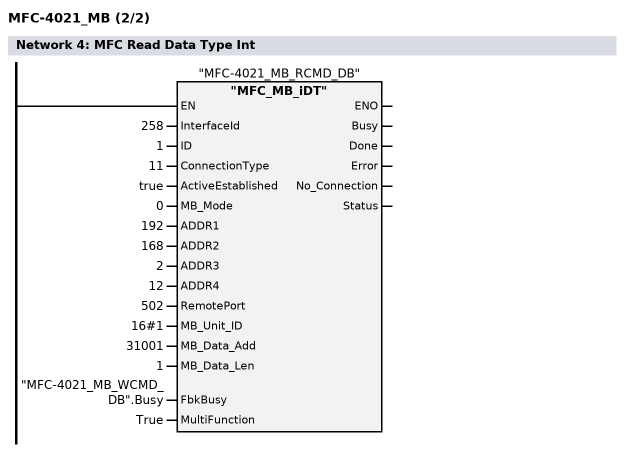
   RUNG wire#powerrail
      "MFC-4021_MB_RCMD_DB"(InterfaceId := 258, ID := 1, ConnectionType := 11, ActiveEstablished := true, MB_Mode := 0, ADDR1 := 192, ADDR2 := 168, ADDR3 := 2, ADDR4 := 12, RemotePort := 502, MB_Unit_ID := 16#1, MB_Data_Add := 31001, MB_Data_Len := 1, FbkBusy := "MFC-4021_MB_WCMD_DB".Busy, MultiFunction := True, Busy =>, Done =>, Error =>, No_Connection =>, Status =>)
   END_RUNG
   // the same network as SCL:
   "MFC-4021_MB_RCMD_DB"(InterfaceId := 258,   // "MFC_MB_iDT"
                         ID := 1,
                         ConnectionType := 11,
                         ActiveEstablished := true,
                         MB_Mode := 0,
                         ADDR1 := 192,
                         ADDR2 := 168,
                         ADDR3 := 2,
                         ADDR4 := 12,
                         RemotePort := 502,
                         MB_Unit_ID := 16#1,
                         MB_Data_Add := 31001,
                         MB_Data_Len := 1,
                         FbkBusy := "MFC-4021_MB_WCMD_DB".Busy,
                         MultiFunction := True);
END_REGION
END_FUNCTION

// folder: Outside Comms/ModBus Comms/MFCs/MFC-4024

FUNCTION "MFC-4024_MB" : Void   // FC78, LAD
{ S7_Optimized_Access := 'TRUE' }
VERSION : 0.1
BEGIN

REGION Network 1: MFC Read Data Type Real
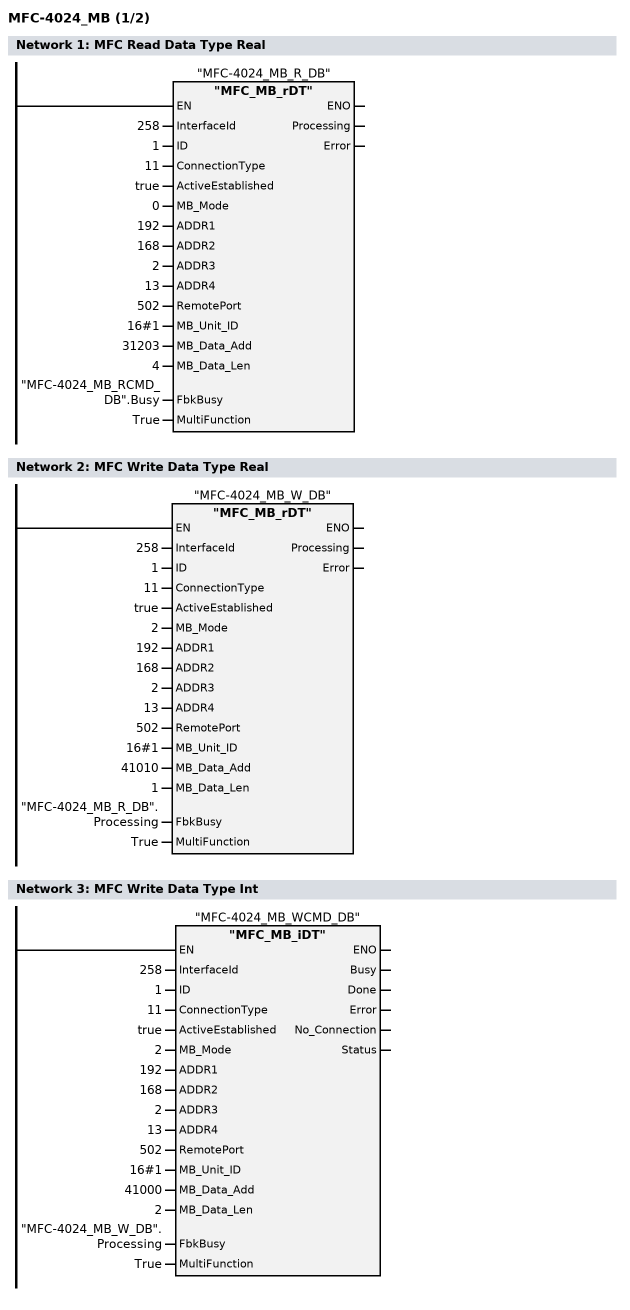
   RUNG wire#powerrail
      "MFC-4024_MB_R_DB"(InterfaceId := 258, ID := 1, ConnectionType := 11, ActiveEstablished := true, MB_Mode := 0, ADDR1 := 192, ADDR2 := 168, ADDR3 := 2, ADDR4 := 13, RemotePort := 502, MB_Unit_ID := 16#1, MB_Data_Add := 31203, MB_Data_Len := 4, FbkBusy := "MFC-4024_MB_RCMD_DB".Busy, MultiFunction := True, Processing =>, Error =>)
   END_RUNG
   // the same network as SCL:
   "MFC-4024_MB_R_DB"(InterfaceId := 258,   // "MFC_MB_rDT"
                      ID := 1,
                      ConnectionType := 11,
                      ActiveEstablished := true,
                      MB_Mode := 0,
                      ADDR1 := 192,
                      ADDR2 := 168,
                      ADDR3 := 2,
                      ADDR4 := 13,
                      RemotePort := 502,
                      MB_Unit_ID := 16#1,
                      MB_Data_Add := 31203,
                      MB_Data_Len := 4,
                      FbkBusy := "MFC-4024_MB_RCMD_DB".Busy,
                      MultiFunction := True);
END_REGION

REGION Network 2: MFC Write Data Type Real
   RUNG wire#powerrail
      "MFC-4024_MB_W_DB"(InterfaceId := 258, ID := 1, ConnectionType := 11, ActiveEstablished := true, MB_Mode := 2, ADDR1 := 192, ADDR2 := 168, ADDR3 := 2, ADDR4 := 13, RemotePort := 502, MB_Unit_ID := 16#1, MB_Data_Add := 41010, MB_Data_Len := 1, FbkBusy := "MFC-4024_MB_R_DB".Processing, MultiFunction := True, Processing =>, Error =>)
   END_RUNG
   // the same network as SCL:
   "MFC-4024_MB_W_DB"(InterfaceId := 258,   // "MFC_MB_rDT"
                      ID := 1,
                      ConnectionType := 11,
                      ActiveEstablished := true,
                      MB_Mode := 2,
                      ADDR1 := 192,
                      ADDR2 := 168,
                      ADDR3 := 2,
                      ADDR4 := 13,
                      RemotePort := 502,
                      MB_Unit_ID := 16#1,
                      MB_Data_Add := 41010,
                      MB_Data_Len := 1,
                      FbkBusy := "MFC-4024_MB_R_DB".Processing,
                      MultiFunction := True);
END_REGION

REGION Network 3: MFC Write Data Type Int
   RUNG wire#powerrail
      "MFC-4024_MB_WCMD_DB"(InterfaceId := 258, ID := 1, ConnectionType := 11, ActiveEstablished := true, MB_Mode := 2, ADDR1 := 192, ADDR2 := 168, ADDR3 := 2, ADDR4 := 13, RemotePort := 502, MB_Unit_ID := 16#1, MB_Data_Add := 41000, MB_Data_Len := 2, FbkBusy := "MFC-4024_MB_W_DB".Processing, MultiFunction := True, Busy =>, Done =>, Error =>, No_Connection =>, Status =>)
   END_RUNG
   // the same network as SCL:
   "MFC-4024_MB_WCMD_DB"(InterfaceId := 258,   // "MFC_MB_iDT"
                         ID := 1,
                         ConnectionType := 11,
                         ActiveEstablished := true,
                         MB_Mode := 2,
                         ADDR1 := 192,
                         ADDR2 := 168,
                         ADDR3 := 2,
                         ADDR4 := 13,
                         RemotePort := 502,
                         MB_Unit_ID := 16#1,
                         MB_Data_Add := 41000,
                         MB_Data_Len := 2,
                         FbkBusy := "MFC-4024_MB_W_DB".Processing,
                         MultiFunction := True);
END_REGION

REGION Network 4: MFC Read Data Type Int
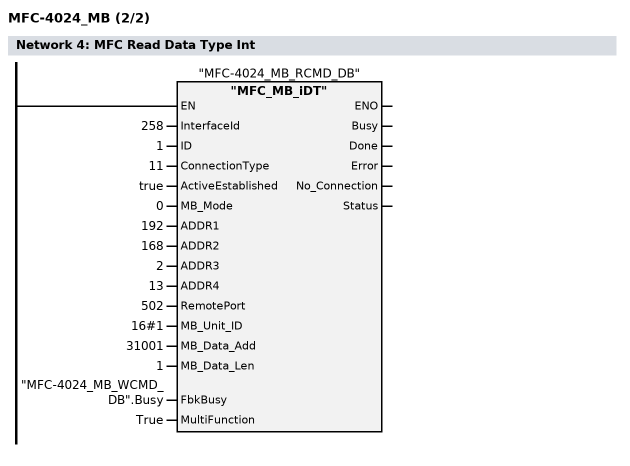
   RUNG wire#powerrail
      "MFC-4024_MB_RCMD_DB"(InterfaceId := 258, ID := 1, ConnectionType := 11, ActiveEstablished := true, MB_Mode := 0, ADDR1 := 192, ADDR2 := 168, ADDR3 := 2, ADDR4 := 13, RemotePort := 502, MB_Unit_ID := 16#1, MB_Data_Add := 31001, MB_Data_Len := 1, FbkBusy := "MFC-4024_MB_WCMD_DB".Busy, MultiFunction := True, Busy =>, Done =>, Error =>, No_Connection =>, Status =>)
   END_RUNG
   // the same network as SCL:
   "MFC-4024_MB_RCMD_DB"(InterfaceId := 258,   // "MFC_MB_iDT"
                         ID := 1,
                         ConnectionType := 11,
                         ActiveEstablished := true,
                         MB_Mode := 0,
                         ADDR1 := 192,
                         ADDR2 := 168,
                         ADDR3 := 2,
                         ADDR4 := 13,
                         RemotePort := 502,
                         MB_Unit_ID := 16#1,
                         MB_Data_Add := 31001,
                         MB_Data_Len := 1,
                         FbkBusy := "MFC-4024_MB_WCMD_DB".Busy,
                         MultiFunction := True);
END_REGION
END_FUNCTION

// folder: Outside Comms/ModBus Comms/MFCs/MFC-4025

FUNCTION "MFC-4025_MB" : Void   // FC93, LAD
{ S7_Optimized_Access := 'TRUE' }
VERSION : 0.1
BEGIN

REGION Network 1: MFC Read Data Type Real
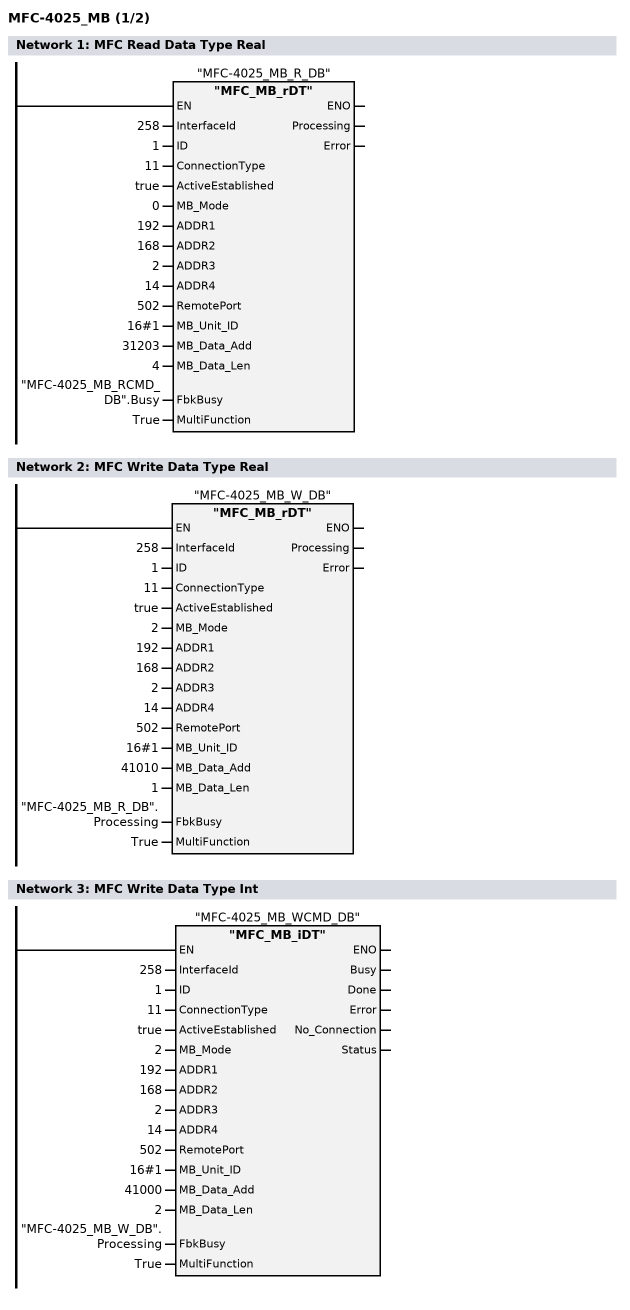
   RUNG wire#powerrail
      "MFC-4025_MB_R_DB"(InterfaceId := 258, ID := 1, ConnectionType := 11, ActiveEstablished := true, MB_Mode := 0, ADDR1 := 192, ADDR2 := 168, ADDR3 := 2, ADDR4 := 14, RemotePort := 502, MB_Unit_ID := 16#1, MB_Data_Add := 31203, MB_Data_Len := 4, FbkBusy := "MFC-4025_MB_RCMD_DB".Busy, MultiFunction := True, Processing =>, Error =>)
   END_RUNG
   // the same network as SCL:
   "MFC-4025_MB_R_DB"(InterfaceId := 258,   // "MFC_MB_rDT"
                      ID := 1,
                      ConnectionType := 11,
                      ActiveEstablished := true,
                      MB_Mode := 0,
                      ADDR1 := 192,
                      ADDR2 := 168,
                      ADDR3 := 2,
                      ADDR4 := 14,
                      RemotePort := 502,
                      MB_Unit_ID := 16#1,
                      MB_Data_Add := 31203,
                      MB_Data_Len := 4,
                      FbkBusy := "MFC-4025_MB_RCMD_DB".Busy,
                      MultiFunction := True);
END_REGION

REGION Network 2: MFC Write Data Type Real
   RUNG wire#powerrail
      "MFC-4025_MB_W_DB"(InterfaceId := 258, ID := 1, ConnectionType := 11, ActiveEstablished := true, MB_Mode := 2, ADDR1 := 192, ADDR2 := 168, ADDR3 := 2, ADDR4 := 14, RemotePort := 502, MB_Unit_ID := 16#1, MB_Data_Add := 41010, MB_Data_Len := 1, FbkBusy := "MFC-4025_MB_R_DB".Processing, MultiFunction := True, Processing =>, Error =>)
   END_RUNG
   // the same network as SCL:
   "MFC-4025_MB_W_DB"(InterfaceId := 258,   // "MFC_MB_rDT"
                      ID := 1,
                      ConnectionType := 11,
                      ActiveEstablished := true,
                      MB_Mode := 2,
                      ADDR1 := 192,
                      ADDR2 := 168,
                      ADDR3 := 2,
                      ADDR4 := 14,
                      RemotePort := 502,
                      MB_Unit_ID := 16#1,
                      MB_Data_Add := 41010,
                      MB_Data_Len := 1,
                      FbkBusy := "MFC-4025_MB_R_DB".Processing,
                      MultiFunction := True);
END_REGION

REGION Network 3: MFC Write Data Type Int
   RUNG wire#powerrail
      "MFC-4025_MB_WCMD_DB"(InterfaceId := 258, ID := 1, ConnectionType := 11, ActiveEstablished := true, MB_Mode := 2, ADDR1 := 192, ADDR2 := 168, ADDR3 := 2, ADDR4 := 14, RemotePort := 502, MB_Unit_ID := 16#1, MB_Data_Add := 41000, MB_Data_Len := 2, FbkBusy := "MFC-4025_MB_W_DB".Processing, MultiFunction := True, Busy =>, Done =>, Error =>, No_Connection =>, Status =>)
   END_RUNG
   // the same network as SCL:
   "MFC-4025_MB_WCMD_DB"(InterfaceId := 258,   // "MFC_MB_iDT"
                         ID := 1,
                         ConnectionType := 11,
                         ActiveEstablished := true,
                         MB_Mode := 2,
                         ADDR1 := 192,
                         ADDR2 := 168,
                         ADDR3 := 2,
                         ADDR4 := 14,
                         RemotePort := 502,
                         MB_Unit_ID := 16#1,
                         MB_Data_Add := 41000,
                         MB_Data_Len := 2,
                         FbkBusy := "MFC-4025_MB_W_DB".Processing,
                         MultiFunction := True);
END_REGION

REGION Network 4: MFC Read Data Type Int
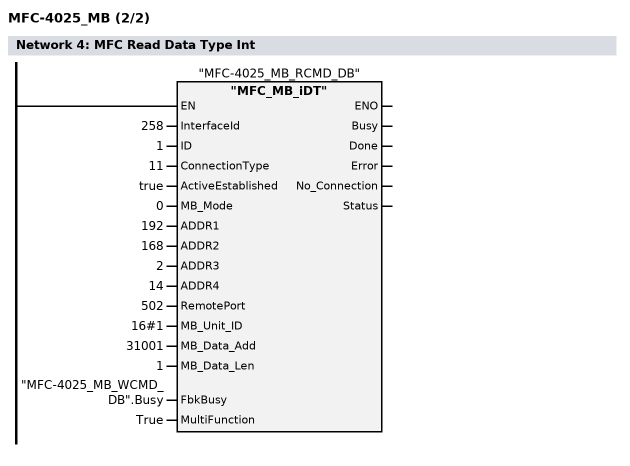
   RUNG wire#powerrail
      "MFC-4025_MB_RCMD_DB"(InterfaceId := 258, ID := 1, ConnectionType := 11, ActiveEstablished := true, MB_Mode := 0, ADDR1 := 192, ADDR2 := 168, ADDR3 := 2, ADDR4 := 14, RemotePort := 502, MB_Unit_ID := 16#1, MB_Data_Add := 31001, MB_Data_Len := 1, FbkBusy := "MFC-4025_MB_WCMD_DB".Busy, MultiFunction := True, Busy =>, Done =>, Error =>, No_Connection =>, Status =>)
   END_RUNG
   // the same network as SCL:
   "MFC-4025_MB_RCMD_DB"(InterfaceId := 258,   // "MFC_MB_iDT"
                         ID := 1,
                         ConnectionType := 11,
                         ActiveEstablished := true,
                         MB_Mode := 0,
                         ADDR1 := 192,
                         ADDR2 := 168,
                         ADDR3 := 2,
                         ADDR4 := 14,
                         RemotePort := 502,
                         MB_Unit_ID := 16#1,
                         MB_Data_Add := 31001,
                         MB_Data_Len := 1,
                         FbkBusy := "MFC-4025_MB_WCMD_DB".Busy,
                         MultiFunction := True);
END_REGION
END_FUNCTION

// folder: Outside Comms/ModBus Comms/pH Transmitters/pH-2011/12

FUNCTION "pH_ModBus" : Void   // FC86, LAD
{ S7_Optimized_Access := 'TRUE' }
VERSION : 0.1
BEGIN

REGION Network 1: pH-2011/12 Modbus Data
   // Collecting pH and Temperatures in real Data Type
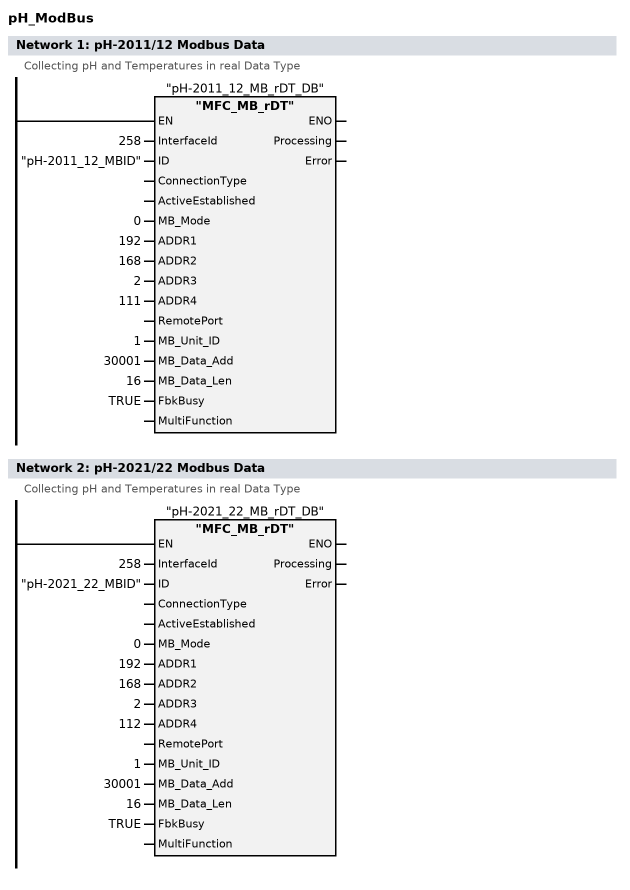
   RUNG wire#powerrail
      "pH-2011_12_MB_rDT_DB"(InterfaceId := 258, ID := "pH-2011_12_MBID", ConnectionType :=, ActiveEstablished :=, MB_Mode := 0, ADDR1 := 192, ADDR2 := 168, ADDR3 := 2, ADDR4 := 111, RemotePort :=, MB_Unit_ID := 1, MB_Data_Add := 30001, MB_Data_Len := 16, FbkBusy := TRUE, MultiFunction :=, Processing =>, Error =>)
   END_RUNG
   // the same network as SCL:
   "pH-2011_12_MB_rDT_DB"(InterfaceId := 258,   // "MFC_MB_rDT"
                          ID := "pH-2011_12_MBID",
                          MB_Mode := 0,
                          ADDR1 := 192,
                          ADDR2 := 168,
                          ADDR3 := 2,
                          ADDR4 := 111,
                          MB_Unit_ID := 1,
                          MB_Data_Add := 30001,
                          MB_Data_Len := 16,
                          FbkBusy := TRUE);
END_REGION

REGION Network 2: pH-2021/22 Modbus Data
   // Collecting pH and Temperatures in real Data Type
   RUNG wire#powerrail
      "pH-2021_22_MB_rDT_DB"(InterfaceId := 258, ID := "pH-2021_22_MBID", ConnectionType :=, ActiveEstablished :=, MB_Mode := 0, ADDR1 := 192, ADDR2 := 168, ADDR3 := 2, ADDR4 := 112, RemotePort :=, MB_Unit_ID := 1, MB_Data_Add := 30001, MB_Data_Len := 16, FbkBusy := TRUE, MultiFunction :=, Processing =>, Error =>)
   END_RUNG
   // the same network as SCL:
   "pH-2021_22_MB_rDT_DB"(InterfaceId := 258,   // "MFC_MB_rDT"
                          ID := "pH-2021_22_MBID",
                          MB_Mode := 0,
                          ADDR1 := 192,
                          ADDR2 := 168,
                          ADDR3 := 2,
                          ADDR4 := 112,
                          MB_Unit_ID := 1,
                          MB_Data_Add := 30001,
                          MB_Data_Len := 16,
                          FbkBusy := TRUE);
END_REGION
END_FUNCTION

// folder: PID Controller

FUNCTION "PIDController" : Void   // FC4, LAD
TITLE = PID Controllers
{ S7_Optimized_Access := 'TRUE' }
VERSION : 0.1
// Location: Cycle_1s OB32
   VAR_TEMP
      "INT" : Int;
      "REAL" : Real;
      INT_1 : Real;
      REAL_1 : Real;
   END_VAR
BEGIN

REGION Network 1: MassFlowControllers
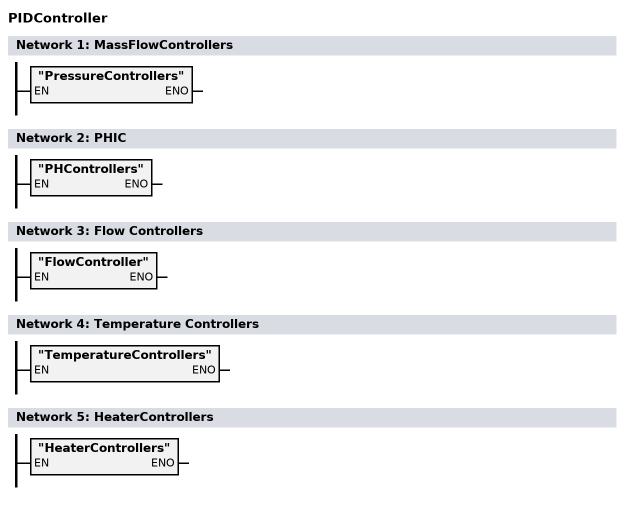
   RUNG wire#powerrail
      "PressureControllers"()
   END_RUNG
   // the same network as SCL:
   "PressureControllers"();
END_REGION

REGION Network 2: PHIC
   RUNG wire#powerrail
      "PHControllers"()
   END_RUNG
   // the same network as SCL:
   "PHControllers"();
END_REGION

REGION Network 3: Flow Controllers
   RUNG wire#powerrail
      "FlowController"()
   END_RUNG
   // the same network as SCL:
   "FlowController"();
END_REGION

REGION Network 4: Temperature Controllers
   RUNG wire#powerrail
      "TemperatureControllers"()
   END_RUNG
   // the same network as SCL:
   "TemperatureControllers"();
END_REGION

REGION Network 5: HeaterControllers
   RUNG wire#powerrail
      "HeaterControllers"()
   END_RUNG
   // the same network as SCL:
   "HeaterControllers"();
END_REGION
END_FUNCTION

// folder: PID Controller/FlowControllers

FUNCTION "FlowController" : Void   // FC22, LAD
{ S7_Optimized_Access := 'TRUE' }
VERSION : 0.1
   VAR_TEMP
      "REAL_R-201" : Real;
      "INT_R-201" : Real;
      "INT_R-202" : Real;
      "REAL_R-202" : Real;
   END_VAR
BEGIN

REGION Network 1: FIC-2011:T-101 to R-201 Flow Controller
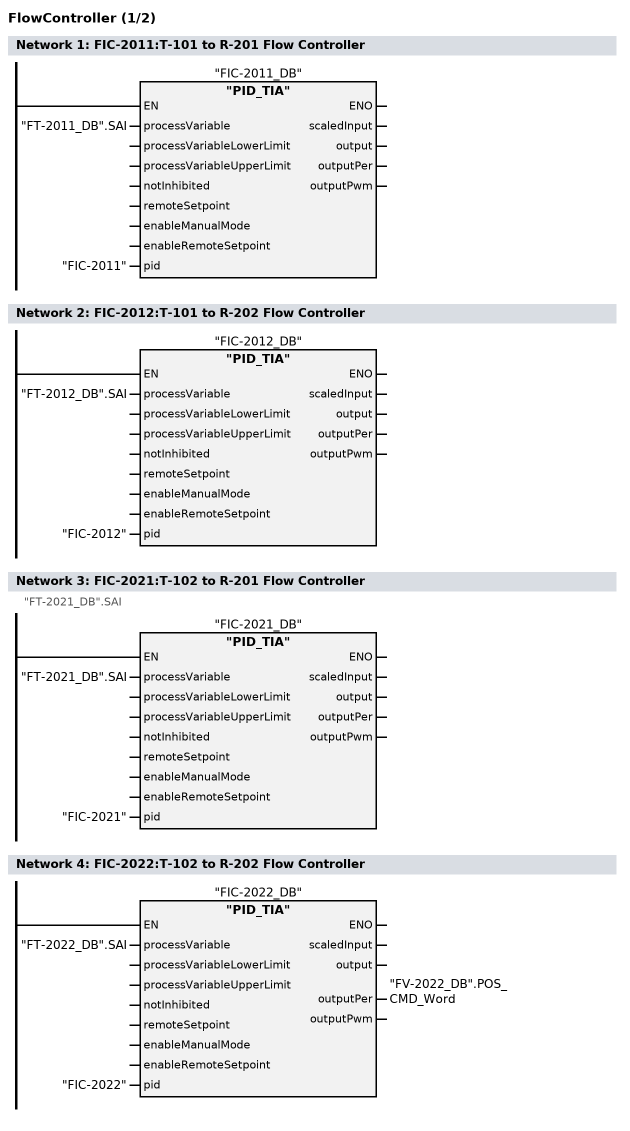
   RUNG wire#powerrail
      "FIC-2011_DB"(processVariable := "FT-2011_DB".SAI, processVariableLowerLimit :=, processVariableUpperLimit :=, notInhibited :=, remoteSetpoint :=, enableManualMode :=, enableRemoteSetpoint :=, pid := "FIC-2011", scaledInput =>, output =>, outputPer =>, outputPwm =>)
   END_RUNG
   // the same network as SCL:
   "FIC-2011_DB"(processVariable := "FT-2011_DB".SAI, pid := "FIC-2011");   // "PID_TIA"
END_REGION

REGION Network 2: FIC-2012:T-101 to R-202 Flow Controller
   RUNG wire#powerrail
      "FIC-2012_DB"(processVariable := "FT-2012_DB".SAI, processVariableLowerLimit :=, processVariableUpperLimit :=, notInhibited :=, remoteSetpoint :=, enableManualMode :=, enableRemoteSetpoint :=, pid := "FIC-2012", scaledInput =>, output =>, outputPer =>, outputPwm =>)
   END_RUNG
   // the same network as SCL:
   "FIC-2012_DB"(processVariable := "FT-2012_DB".SAI, pid := "FIC-2012");   // "PID_TIA"
END_REGION

REGION Network 3: FIC-2021:T-102 to R-201 Flow Controller
   // "FT-2021_DB".SAI
   RUNG wire#powerrail
      "FIC-2021_DB"(processVariable := "FT-2021_DB".SAI, processVariableLowerLimit :=, processVariableUpperLimit :=, notInhibited :=, remoteSetpoint :=, enableManualMode :=, enableRemoteSetpoint :=, pid := "FIC-2021", scaledInput =>, output =>, outputPer =>, outputPwm =>)
   END_RUNG
   // the same network as SCL:
   "FIC-2021_DB"(processVariable := "FT-2021_DB".SAI, pid := "FIC-2021");   // "PID_TIA"
END_REGION

REGION Network 4: FIC-2022:T-102 to R-202 Flow Controller
   RUNG wire#powerrail
      "FIC-2022_DB"(processVariable := "FT-2022_DB".SAI, processVariableLowerLimit :=, processVariableUpperLimit :=, notInhibited :=, remoteSetpoint :=, enableManualMode :=, enableRemoteSetpoint :=, pid := "FIC-2022", scaledInput =>, output =>, outputPer => "FV-2022_DB".POS_CMD_Word, outputPwm =>)
   END_RUNG
   // the same network as SCL:
   "FIC-2022_DB"(processVariable := "FT-2022_DB".SAI, pid := "FIC-2022", outputPer => "FV-2022_DB".POS_CMD_Word);   // "PID_TIA"
END_REGION

REGION Network 5: FIC-3011: Centrifuge Flow Controller
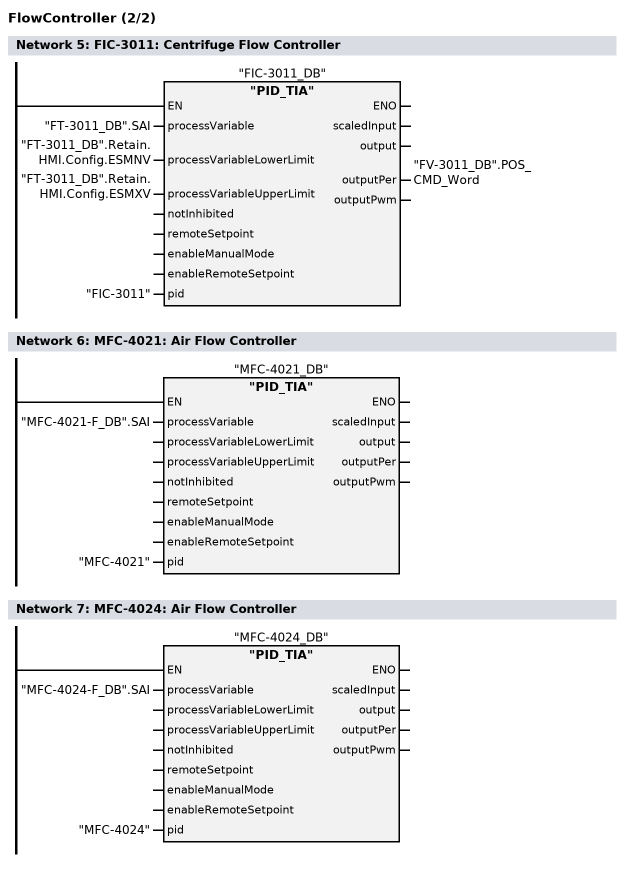
   RUNG wire#powerrail
      "FIC-3011_DB"(processVariable := "FT-3011_DB".SAI, processVariableLowerLimit := "FT-3011_DB".Retain.HMI.Config.ESMNV, processVariableUpperLimit := "FT-3011_DB".Retain.HMI.Config.ESMXV, notInhibited :=, remoteSetpoint :=, enableManualMode :=, enableRemoteSetpoint :=, pid := "FIC-3011", scaledInput =>, output =>, outputPer => "FV-3011_DB".POS_CMD_Word, outputPwm =>)
   END_RUNG
   // the same network as SCL:
   "FIC-3011_DB"(processVariable := "FT-3011_DB".SAI,   // "PID_TIA"
                 processVariableLowerLimit := "FT-3011_DB".Retain.HMI.Config.ESMNV,
                 processVariableUpperLimit := "FT-3011_DB".Retain.HMI.Config.ESMXV,
                 pid := "FIC-3011",
                 outputPer => "FV-3011_DB".POS_CMD_Word);
END_REGION

REGION Network 6: MFC-4021: Air Flow Controller
   RUNG wire#powerrail
      "MFC-4021_DB"(processVariable := "MFC-4021-F_DB".SAI, processVariableLowerLimit :=, processVariableUpperLimit :=, notInhibited :=, remoteSetpoint :=, enableManualMode :=, enableRemoteSetpoint :=, pid := "MFC-4021", scaledInput =>, output =>, outputPer =>, outputPwm =>)
   END_RUNG
   // the same network as SCL:
   "MFC-4021_DB"(processVariable := "MFC-4021-F_DB".SAI, pid := "MFC-4021");   // "PID_TIA"
END_REGION

REGION Network 7: MFC-4024: Air Flow Controller
   RUNG wire#powerrail
      "MFC-4024_DB"(processVariable := "MFC-4024-F_DB".SAI, processVariableLowerLimit :=, processVariableUpperLimit :=, notInhibited :=, remoteSetpoint :=, enableManualMode :=, enableRemoteSetpoint :=, pid := "MFC-4024", scaledInput =>, output =>, outputPer =>, outputPwm =>)
   END_RUNG
   // the same network as SCL:
   "MFC-4024_DB"(processVariable := "MFC-4024-F_DB".SAI, pid := "MFC-4024");   // "PID_TIA"
END_REGION
END_FUNCTION

// folder: PID Controller/Heater Controllers

FUNCTION "HeaterControllers" : Void   // FC27, LAD
{ S7_Optimized_Access := 'TRUE' }
VERSION : 0.1
BEGIN

REGION Network 1: HFC-201
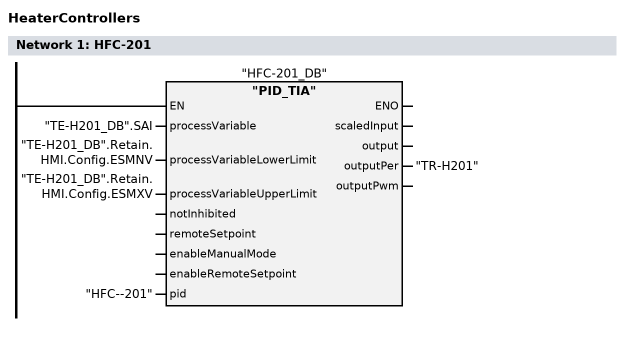
   RUNG wire#powerrail
      "HFC-201_DB"(processVariable := "TE-H201_DB".SAI, processVariableLowerLimit := "TE-H201_DB".Retain.HMI.Config.ESMNV, processVariableUpperLimit := "TE-H201_DB".Retain.HMI.Config.ESMXV, notInhibited :=, remoteSetpoint :=, enableManualMode :=, enableRemoteSetpoint :=, pid := "HFC--201", scaledInput =>, output =>, outputPer => "TR-H201", outputPwm =>)
   END_RUNG
   // the same network as SCL:
   "HFC-201_DB"(processVariable := "TE-H201_DB".SAI,   // "PID_TIA"
                processVariableLowerLimit := "TE-H201_DB".Retain.HMI.Config.ESMNV,
                processVariableUpperLimit := "TE-H201_DB".Retain.HMI.Config.ESMXV,
                pid := "HFC--201",
                outputPer => "TR-H201");
END_REGION
END_FUNCTION

// folder: PID Controller/Level Controllers

FUNCTION "LevelControllers" : Void   // FC21, LAD
{ S7_Optimized_Access := 'TRUE' }
VERSION : 0.1
   VAR_TEMP
      IN : Bool;
      OUT : Bool;
      TRIGGER : Bool;
   END_VAR
   VAR CONSTANT
      MANUAL : Int := 4;
      REMOTE : Int := 6;
   END_VAR
BEGIN
END_FUNCTION

// folder: PID Controller/PH Controllers

FUNCTION "PHControllers" : Void   // FC23, LAD
{ S7_Optimized_Access := 'TRUE' }
VERSION : 0.1
BEGIN

REGION Network 1: PHIC-R-201: R-201 Reactor PH Controller
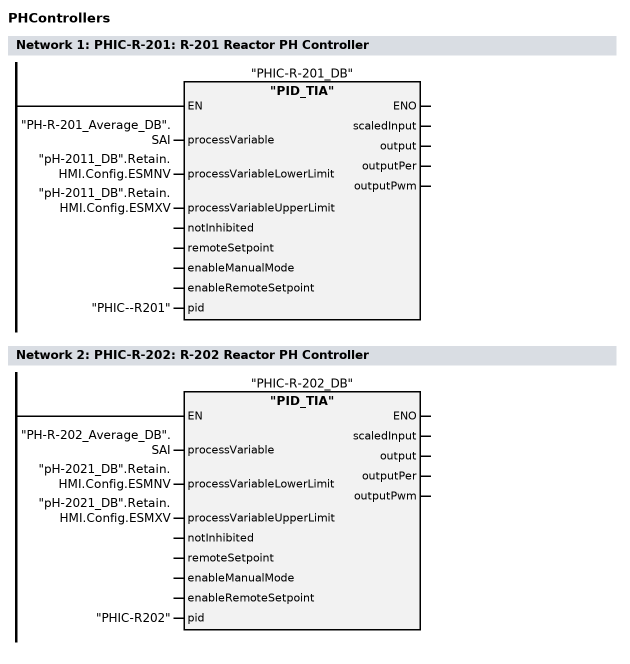
   RUNG wire#powerrail
      "PHIC-R-201_DB"(processVariable := "PH-R-201_Average_DB".SAI, processVariableLowerLimit := "pH-2011_DB".Retain.HMI.Config.ESMNV, processVariableUpperLimit := "pH-2011_DB".Retain.HMI.Config.ESMXV, notInhibited :=, remoteSetpoint :=, enableManualMode :=, enableRemoteSetpoint :=, pid := "PHIC--R201", scaledInput =>, output =>, outputPer =>, outputPwm =>)
   END_RUNG
   // the same network as SCL:
   "PHIC-R-201_DB"(processVariable := "PH-R-201_Average_DB".SAI,   // "PID_TIA"
                   processVariableLowerLimit := "pH-2011_DB".Retain.HMI.Config.ESMNV,
                   processVariableUpperLimit := "pH-2011_DB".Retain.HMI.Config.ESMXV,
                   pid := "PHIC--R201");
END_REGION

REGION Network 2: PHIC-R-202: R-202 Reactor PH Controller
   RUNG wire#powerrail
      "PHIC-R-202_DB"(processVariable := "PH-R-202_Average_DB".SAI, processVariableLowerLimit := "pH-2021_DB".Retain.HMI.Config.ESMNV, processVariableUpperLimit := "pH-2021_DB".Retain.HMI.Config.ESMXV, notInhibited :=, remoteSetpoint :=, enableManualMode :=, enableRemoteSetpoint :=, pid := "PHIC-R202", scaledInput =>, output =>, outputPer =>, outputPwm =>)
   END_RUNG
   // the same network as SCL:
   "PHIC-R-202_DB"(processVariable := "PH-R-202_Average_DB".SAI,   // "PID_TIA"
                   processVariableLowerLimit := "pH-2021_DB".Retain.HMI.Config.ESMNV,
                   processVariableUpperLimit := "pH-2021_DB".Retain.HMI.Config.ESMXV,
                   pid := "PHIC-R202");
END_REGION
END_FUNCTION

// folder: PID Controller/PressureControllers

FUNCTION "PressureControllers" : Void   // FC24, LAD
{ S7_Optimized_Access := 'TRUE' }
VERSION : 0.1
BEGIN

REGION Network 1: MFC-4011 (Air ALICAT to Calcination Furnace R-401)
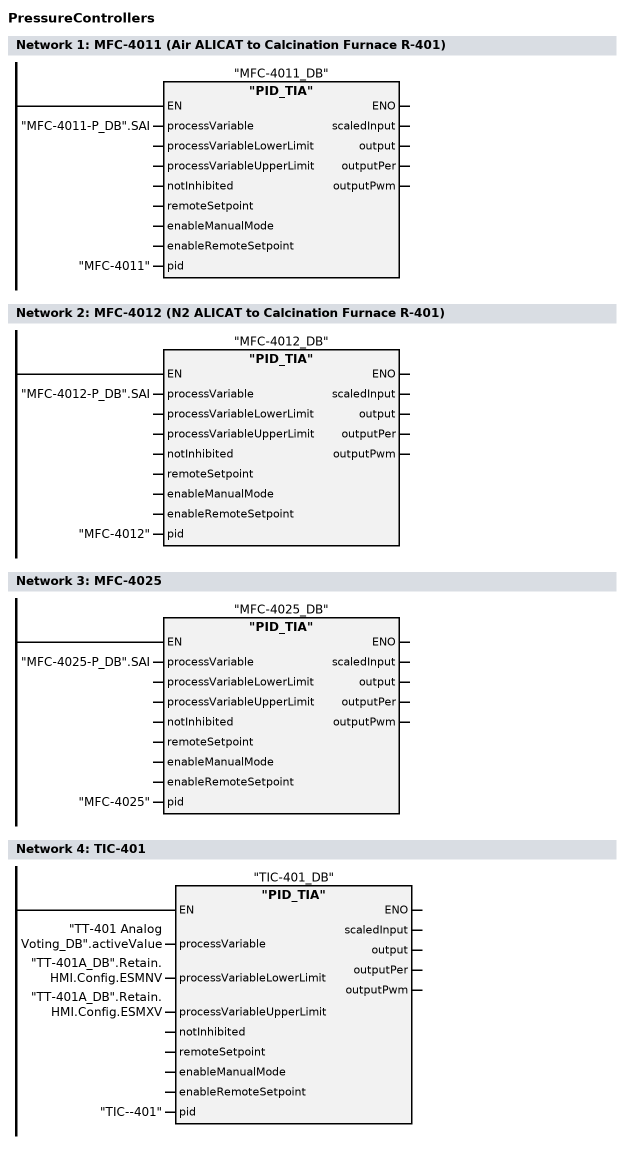
   RUNG wire#powerrail
      "MFC-4011_DB"(processVariable := "MFC-4011-P_DB".SAI, processVariableLowerLimit :=, processVariableUpperLimit :=, notInhibited :=, remoteSetpoint :=, enableManualMode :=, enableRemoteSetpoint :=, pid := "MFC-4011", scaledInput =>, output =>, outputPer =>, outputPwm =>)
   END_RUNG
   // the same network as SCL:
   "MFC-4011_DB"(processVariable := "MFC-4011-P_DB".SAI, pid := "MFC-4011");   // "PID_TIA"
END_REGION

REGION Network 2: MFC-4012 (N2 ALICAT to Calcination Furnace R-401)
   RUNG wire#powerrail
      "MFC-4012_DB"(processVariable := "MFC-4012-P_DB".SAI, processVariableLowerLimit :=, processVariableUpperLimit :=, notInhibited :=, remoteSetpoint :=, enableManualMode :=, enableRemoteSetpoint :=, pid := "MFC-4012", scaledInput =>, output =>, outputPer =>, outputPwm =>)
   END_RUNG
   // the same network as SCL:
   "MFC-4012_DB"(processVariable := "MFC-4012-P_DB".SAI, pid := "MFC-4012");   // "PID_TIA"
END_REGION

REGION Network 3: MFC-4025
   RUNG wire#powerrail
      "MFC-4025_DB"(processVariable := "MFC-4025-P_DB".SAI, processVariableLowerLimit :=, processVariableUpperLimit :=, notInhibited :=, remoteSetpoint :=, enableManualMode :=, enableRemoteSetpoint :=, pid := "MFC-4025", scaledInput =>, output =>, outputPer =>, outputPwm =>)
   END_RUNG
   // the same network as SCL:
   "MFC-4025_DB"(processVariable := "MFC-4025-P_DB".SAI, pid := "MFC-4025");   // "PID_TIA"
END_REGION

REGION Network 4: TIC-401
   RUNG wire#powerrail
      "TIC-401_DB"(processVariable := "TT-401 Analog Voting_DB".activeValue, processVariableLowerLimit := "TT-401A_DB".Retain.HMI.Config.ESMNV, processVariableUpperLimit := "TT-401A_DB".Retain.HMI.Config.ESMXV, notInhibited :=, remoteSetpoint :=, enableManualMode :=, enableRemoteSetpoint :=, pid := "TIC--401", scaledInput =>, output =>, outputPer =>, outputPwm =>)
   END_RUNG
   // the same network as SCL:
   "TIC-401_DB"(processVariable := "TT-401 Analog Voting_DB".activeValue,   // "PID_TIA"
                processVariableLowerLimit := "TT-401A_DB".Retain.HMI.Config.ESMNV,
                processVariableUpperLimit := "TT-401A_DB".Retain.HMI.Config.ESMXV,
                pid := "TIC--401");
END_REGION
END_FUNCTION

// folder: PID Controller/Temperature Controllers

FUNCTION "TemperatureControllers" : Void   // FC26, LAD
{ S7_Optimized_Access := 'TRUE' }
VERSION : 0.1
BEGIN

REGION Network 1: TIC-402A : Zone A Controller
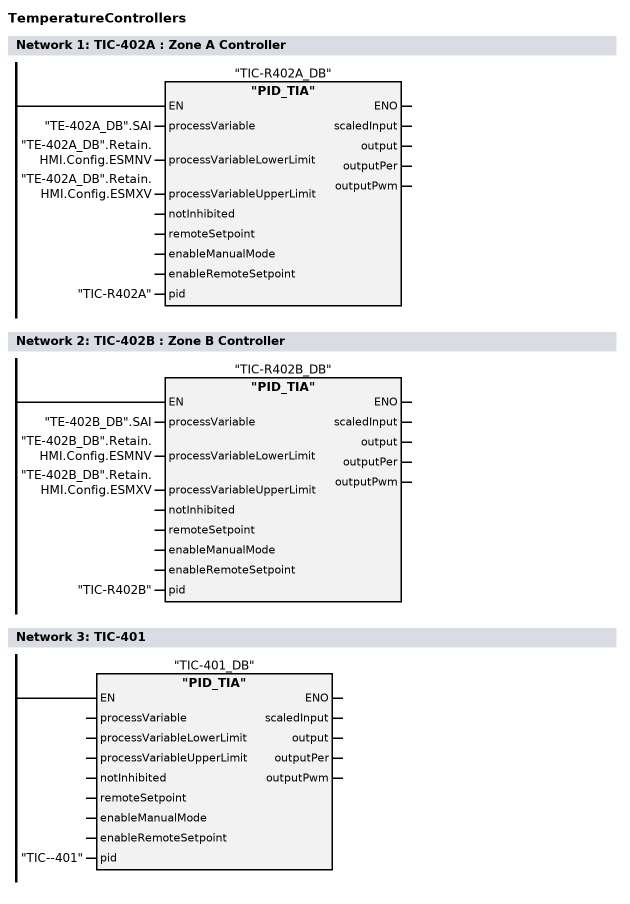
   RUNG wire#powerrail
      "TIC-R402A_DB"(processVariable := "TE-402A_DB".SAI, processVariableLowerLimit := "TE-402A_DB".Retain.HMI.Config.ESMNV, processVariableUpperLimit := "TE-402A_DB".Retain.HMI.Config.ESMXV, notInhibited :=, remoteSetpoint :=, enableManualMode :=, enableRemoteSetpoint :=, pid := "TIC-R402A", scaledInput =>, output =>, outputPer =>, outputPwm =>)
   END_RUNG
   // the same network as SCL:
   "TIC-R402A_DB"(processVariable := "TE-402A_DB".SAI,   // "PID_TIA"
                  processVariableLowerLimit := "TE-402A_DB".Retain.HMI.Config.ESMNV,
                  processVariableUpperLimit := "TE-402A_DB".Retain.HMI.Config.ESMXV,
                  pid := "TIC-R402A");
END_REGION

REGION Network 2: TIC-402B : Zone B Controller
   RUNG wire#powerrail
      "TIC-R402B_DB"(processVariable := "TE-402B_DB".SAI, processVariableLowerLimit := "TE-402B_DB".Retain.HMI.Config.ESMNV, processVariableUpperLimit := "TE-402B_DB".Retain.HMI.Config.ESMXV, notInhibited :=, remoteSetpoint :=, enableManualMode :=, enableRemoteSetpoint :=, pid := "TIC-R402B", scaledInput =>, output =>, outputPer =>, outputPwm =>)
   END_RUNG
   // the same network as SCL:
   "TIC-R402B_DB"(processVariable := "TE-402B_DB".SAI,   // "PID_TIA"
                  processVariableLowerLimit := "TE-402B_DB".Retain.HMI.Config.ESMNV,
                  processVariableUpperLimit := "TE-402B_DB".Retain.HMI.Config.ESMXV,
                  pid := "TIC-R402B");
END_REGION

REGION Network 3: TIC-401
   RUNG wire#powerrail
      "TIC-401_DB"(processVariable :=, processVariableLowerLimit :=, processVariableUpperLimit :=, notInhibited :=, remoteSetpoint :=, enableManualMode :=, enableRemoteSetpoint :=, pid := "TIC--401", scaledInput =>, output =>, outputPer =>, outputPwm =>)
   END_RUNG
   // the same network as SCL:
   "TIC-401_DB"(pid := "TIC--401");   // "PID_TIA"
END_REGION
END_FUNCTION

// folder: Pumps

FUNCTION "Simple_Pump" : Void   // FC9, LAD
{ S7_Optimized_Access := 'TRUE' }
VERSION : 0.1
   VAR_TEMP
      PMP_TIMEOUT : Bool;
      PMP_TIMEOUT_TIME : Time;
      ON : Bool;
   END_VAR
BEGIN

REGION Network 1 (SCL): p-104 interlock Senario
   (*IF "XV-1041_DB".CS AND "XV-1042_DB".CS AND "XV-1043_DB".CS AND "XV-1044_DB".CS AND "P-104A_DB".CF OR "P-104B_DB".CF = TRUE THEN
       #ON := TRUE;
       "P-104_Run_timeout".TON(IN := #ON,
                              PT := T#10s,
                              Q => #PMP_TIMEOUT,
                               ET => #PMP_TIMEOUT_TIME);
       IF #PMP_TIMEOUT = TRUE THEN
          "P-104A_DB".IL := FALSE;
          "P-104A_DB".ON := FALSE;
          "P-104A_DB".HMI.Controls.Start := FALSE;
          "P-104A_DB".OFF := TRUE;
         "P-104A_DB".HMI.Controls.Stop := TRUE;
          "P-104B_DB".IL := FALSE;
         "P-104B_DB".ON := FALSE;
         "P-104B_DB".HMI.Controls.Start := FALSE;
          "P-104B_DB".OFF := TRUE;
          "P-104B_DB".HMI.Controls.Stop := TRUE;
     END_IF;

   ELSE
       "P-104A_DB".IL:= TRUE;
      "P-104B_DB".IL:= TRUE;
     #ON := FALSE;
      #PMP_TIMEOUT := FALSE;
      RESET_TIMER("P-104_Run_timeout");
   END_IF;*)
END_REGION

REGION Network 2: P-104A